// TIA Portal project "OP-TQ-01" (V13)

(* hardware
DEVICE "S7-1200 station_1"  S7-1200 Station
   slot 0: "Rack_0"  Rack  V1.0
   slot 1: "PLC_1"  CPU 1214C DC/DC/Rly  6ES7 214-1HG31-0XB0  V3.0
   slot 2: "AI 4x13BIT_1"  6ES7 231-4HD30-0XB0  V1.0
   slot 3: "AI 4x13BIT_2"  6ES7 231-4HD30-0XB0  V1.0
   slot 4: "AQ 2x14BIT_1"  6ES7 232-4HB32-0XB0  V2.0
DEVICE "HMI_1"  KP400 Comfort
   slot 0: "HMI"  HMI  6AV2 124-1DC01-0AX0  13.0.1.0
   slot 1: "HMI_RT_1"  KP400 Comfort  6AV2 124-1DC01-0AX0  13.0.1.0
   slot 5: "HMI_1.IE_CP_1"  PROFINET Interface
      slot 1: "PROFINET Interface_1"  PROFINET Interface
         slot 1: "Port_1"  Port
   slot 7: "HMI_1.MPI/DP_CP_1"  MPI/DP Interface
*)

// ===== PLC "PLC_1"  CPU 1214C DC/DC/Rly =====

VAR_GLOBAL   // PLC tag table "Default tag table"
   "System_Byte" AT %MB1 : Byte;
   "FirstScan" AT %M1.0 : Bool;
   "DiagStatusUpdate" AT %M1.1 : Bool;
   "AlwaysTRUE" AT %M1.2 : Bool;
   "AlwaysFALSE" AT %M1.3 : Bool;
   "Clock_Byte" AT %MB0 : Byte;
   "Clock_10Hz" AT %M0.0 : Bool;
   "Clock_5Hz" AT %M0.1 : Bool;
   "Clock_2.5Hz" AT %M0.2 : Bool;
   "Clock_2Hz" AT %M0.3 : Bool;
   "Clock_1.25Hz" AT %M0.4 : Bool;
   "Clock_1Hz" AT %M0.5 : Bool;
   "Clock_0.625Hz" AT %M0.6 : Bool;
   "Clock_0.5Hz" AT %M0.7 : Bool;
   "TT-006-EA" AT %IW96 : Int;
   "TT-007-EA" AT %IW98 : Int;
   "TT-008-EA" AT %IW100 : Int;
   "TT-009-EA" AT %IW102 : Int;
   "TT-010-EA" AT %IW104 : Int;
   "TT-011-EA" AT %IW106 : Int;
   "LT-009-EA" AT %IW108 : Int;
   "LT-CX-REC-EA" AT %IW110 : Int;
   "LSLL-004" AT %I0.0 : Bool;
   "TSH-004" AT %I0.1 : Bool;
   "TERMICO" AT %I0.2 : Bool;
   "RESISTENCIAS-MAN-AUTO" AT %I0.3 : Bool;
   "RESISTENCIAS-RETORNO" AT %I0.4 : Bool;
   "BOTAO-LIGA" AT %I0.5 : Bool;
   "BOTAO-DESLIGA" AT %I0.6 : Bool;
   "FALTA-DE-FASE" AT %I0.7 : Bool;
   "RESISTENCIAS-DESLIGA" AT %Q0.0 : Bool;
   "R2-DESLIGA" AT %Q0.1 : Bool;
   "CX-REC-NIVEL-H" AT %Q0.2 : Bool;
   "CX-REC-NIVEL-HH" AT %Q0.3 : Bool;
   "AlarmAnalog" AT %M13.0 : Bool;
   "REC_ALM" AT %M2.0 : Bool;
   "IW0" AT %IW0 : Word;
   "SAIDAS_DIGITAIS" AT %QW0 : Word;
   "R01A-Liga" AT %M110.0 : Bool;
   "R01B-Liga" AT %M110.1 : Bool;
   "R01C-Liga" AT %M110.2 : Bool;
   "R01D-Liga" AT %M110.3 : Bool;
   "R01E-Liga" AT %M110.4 : Bool;
   "R01F-Liga" AT %M110.5 : Bool;
   "Intlok-Resist" AT %M110.6 : Bool;
   "Tag_1" AT %MW140 : Int;
   "Tag_2" AT %MW142 : Int;
   "Tag_3" AT %MW144 : Int;
   "Tag_4" AT %M20.0 : Bool;
   "Tag_5" AT %M20.1 : Bool;
END_VAR

TYPE "Alm-Bits"
   STRUCT
      UDF : Bool;
      UDR : Bool;
      OVF : Bool;
      OVR : Bool;
      HH : Bool;
      H : Bool;
      L : Bool;
      LL : Bool;
   END_STRUCT;
END_TYPE

TYPE "SP-Temperaturas"
   STRUCT
      AuxLiga : Bool;
      ErroSP : Bool;
      "SP-MAX" : Real;
      "SP-MIN" : Real;
   END_STRUCT;
END_TYPE

// folder: 0000 - AUXILIARES

DATA_BLOCK "TIMERS"   // DB5100
{ S7_Optimized_Access := 'FALSE' }
VERSION : 0.1
   VAR
      T : Array[0..25] of IEC_TIMER;
   END_VAR
BEGIN
END_DATA_BLOCK

// folder: 0020 - ENTRADAS DIGITAIS

DATA_BLOCK "ED"   // DB20
TITLE = ESPELHO DAS ENTRADAS DIGITAIS
{ S7_Optimized_Access := 'FALSE' }
VERSION : 0.1
   VAR
      "LSLL-004" : Bool;
      "TSH-004" : Bool;
      TERMICO : Bool;
      "RESISTENCIAS-LOC-REM" : Bool;
      "RESISTENCIAS-RETORNO" : Bool;
      "BOTAO-LIGA" : Bool;
      "BOTAO-DESLIGA" : Bool;
      "FALTA-DE-FASE" : Bool;
      RESERVA_1 : Bool;
      RESERVA_2 : Bool;
      RESERVA_3 : Bool;
      RESERVA_4 : Bool;
      RESERVA_5 : Bool;
      RESERVA_6 : Bool;
      RESERVA_7 : Bool;
      RESERVA_8 : Bool;
      RESERVA : Array[2..3] of Byte;
   END_VAR
BEGIN
END_DATA_BLOCK

// folder: 0030 - SAIDAS DIGITAIS

DATA_BLOCK "SD"   // DB30
TITLE = ESPELHO DAS SAÍDAS DIGITAIS
{ S7_Optimized_Access := 'FALSE' }
VERSION : 0.1
   VAR
      "LD-RESISTENCIAS" : Bool;
      "R2-DESLIGA" : Bool;
      "CX-REC-NIVEL-H" : Bool;
      "CX-REC-NIVEL-HH" : Bool;
      RESERVA_1 : Bool;
      RESERVA_2 : Bool;
      RESERVA_3 : Bool;
      RESERVA_4 : Bool;
      RESERVA_5 : Bool;
      RESERVA_6 : Bool;
      RESERVA_7 : Bool;
      RESERVA_8 : Bool;
      RESERVA_9 : Bool;
      RESERVA_10 : Bool;
      RESERVA_11 : Bool;
      RESERVA_12 : Bool;
      RESERVA : Array[2..3] of Byte;
   END_VAR
BEGIN
END_DATA_BLOCK

// folder: 1100 - ACIONAMENTOS/RESISTENCIAS

DATA_BLOCK "R01A-R01F"   // DB1101
{ S7_Optimized_Access := 'FALSE' }
VERSION : 0.1
// stored: InstanceOfName 1110 - RESISTENCIAS
"1110 - RESISTENCIAS"
BEGIN
END_DATA_BLOCK

DATA_BLOCK "SP-TT"   // DB1110
{ S7_Optimized_Access := 'FALSE' }
VERSION : 0.1
   VAR
      "TT-006-R01A" : "SP-Temperaturas";
      "TT-007-R01B" : "SP-Temperaturas";
      "TT-008-R01C" : "SP-Temperaturas";
      "TT-009-R01D" : "SP-Temperaturas";
      "TT-010-R01E" : "SP-Temperaturas";
      "TT-011-R01F" : "SP-Temperaturas";
   END_VAR
BEGIN
END_DATA_BLOCK

// folder: 1300 - ALARMES

DATA_BLOCK "ALM"   // DB1301
{ S7_Optimized_Access := 'FALSE' }
VERSION : 0.1
   VAR
      "LSLL-004" : Bool;
      "TSH-004" : Bool;
      FaltaDeFase : Bool;
      RESERVA : Word;
   END_VAR
BEGIN
END_DATA_BLOCK

// folder: 1400 - ENTRADAS ANALOGICAS/NIVEL

DATA_BLOCK "LT-009"   // DB1417
{ S7_Optimized_Access := 'FALSE' }
VERSION : 0.1
// stored: InstanceOfName 1401 - LEITURAS ANALÓGICAS 1HAB
"1401 - LEITURAS ANALÓGICAS 1HAB"
BEGIN
END_DATA_BLOCK

DATA_BLOCK "LT-008"   // DB1418
{ S7_Optimized_Access := 'FALSE' }
VERSION : 0.1
// stored: InstanceOfName 1401 - LEITURAS ANALÓGICAS 1HAB
"1401 - LEITURAS ANALÓGICAS 1HAB"
BEGIN
END_DATA_BLOCK

// folder: 1400 - ENTRADAS ANALOGICAS/TEMPERATURA

DATA_BLOCK "TT-006-R01A"   // DB1411
{ S7_Optimized_Access := 'FALSE' }
VERSION : 0.1
// stored: InstanceOfName 1401 - LEITURAS ANALÓGICAS 1HAB
"1401 - LEITURAS ANALÓGICAS 1HAB"
BEGIN
END_DATA_BLOCK

DATA_BLOCK "TT-007-R01B"   // DB1412
{ S7_Optimized_Access := 'FALSE' }
VERSION : 0.1
// stored: InstanceOfName 1401 - LEITURAS ANALÓGICAS 1HAB
"1401 - LEITURAS ANALÓGICAS 1HAB"
BEGIN
END_DATA_BLOCK

DATA_BLOCK "TT-008-R01C"   // DB1413
{ S7_Optimized_Access := 'FALSE' }
VERSION : 0.1
// stored: InstanceOfName 1401 - LEITURAS ANALÓGICAS 1HAB
"1401 - LEITURAS ANALÓGICAS 1HAB"
BEGIN
END_DATA_BLOCK

DATA_BLOCK "TT-009-R01D"   // DB1414
{ S7_Optimized_Access := 'FALSE' }
VERSION : 0.1
// stored: InstanceOfName 1401 - LEITURAS ANALÓGICAS 1HAB
"1401 - LEITURAS ANALÓGICAS 1HAB"
BEGIN
END_DATA_BLOCK

DATA_BLOCK "TT-010-R01E"   // DB1415
{ S7_Optimized_Access := 'FALSE' }
VERSION : 0.1
// stored: InstanceOfName 1401 - LEITURAS ANALÓGICAS 1HAB
"1401 - LEITURAS ANALÓGICAS 1HAB"
BEGIN
END_DATA_BLOCK

DATA_BLOCK "TT-011-R01F"   // DB1416
{ S7_Optimized_Access := 'FALSE' }
VERSION : 0.1
// stored: InstanceOfName 1401 - LEITURAS ANALÓGICAS 1HAB
"1401 - LEITURAS ANALÓGICAS 1HAB"
BEGIN
END_DATA_BLOCK

// folder: (top level)

ORGANIZATION_BLOCK "Main"   // OB1, LAD, ProgramCycle
TITLE = "Main Program Sweep (Cycle)"
{ S7_Optimized_Access := 'FALSE' }
VERSION : 0.1
BEGIN

REGION Network 1
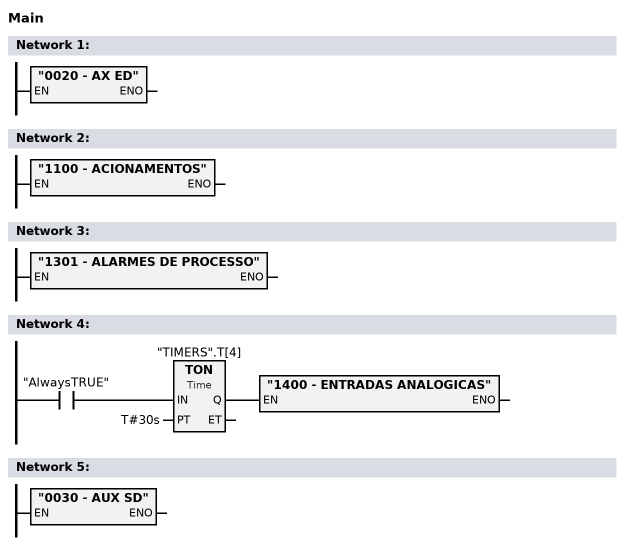
   RUNG wire#powerrail
      "0020 - AX ED"()
   END_RUNG
   // the same network as SCL:
   "0020 - AX ED"();
END_REGION

REGION Network 2
   RUNG wire#powerrail
      "1100 - ACIONAMENTOS"()
   END_RUNG
   // the same network as SCL:
   "1100 - ACIONAMENTOS"();
END_REGION

REGION Network 3
   RUNG wire#powerrail
      "1301 - ALARMES DE PROCESSO"()
   END_RUNG
   // the same network as SCL:
   "1301 - ALARMES DE PROCESSO"();
END_REGION

REGION Network 4
   "TIMERS".T[4].TON(IN := "AlwaysTRUE", PT := T#30s);
   IF "TIMERS".T[4].Q THEN "1400 - ENTRADAS ANALOGICAS"(); END_IF;
END_REGION

REGION Network 5
   RUNG wire#powerrail
      "0030 - AUX SD"()
   END_RUNG
   // the same network as SCL:
   "0030 - AUX SD"();
END_REGION
END_ORGANIZATION_BLOCK

// folder: 0020 - ENTRADAS DIGITAIS

FUNCTION "0020 - AX ED" : Void   // FC20, LAD
TITLE = ESPELHO DAS ENTRADAS DIGITAIS
{ S7_Optimized_Access := 'FALSE' }
VERSION : 0.1
BEGIN

REGION Network 1: ESPELHA AS ENTRADAS DIGITAIS DO CLP
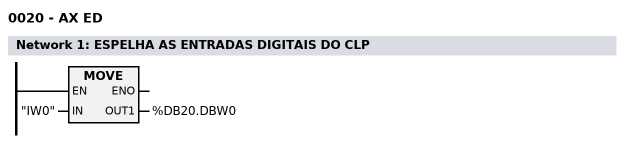
   RUNG wire#powerrail
      { S7_GenerateENO := "TRUE" } Move(in := "IW0", out1 => %DB20.DBW0)
   END_RUNG
   // the same network as SCL:
   %DB20.DBW0 := "IW0";
END_REGION
END_FUNCTION

// folder: 0030 - SAIDAS DIGITAIS

FUNCTION "0030 - AUX SD" : Void   // FC30, LAD
TITLE = ESPELHO DAS SAIDAS DIGITAIS
{ S7_Optimized_Access := 'FALSE' }
VERSION : 0.1
BEGIN

REGION Network 1: ESPELHO DAS SAIDAS DIGITAIS DAS ECP1 E ECP2
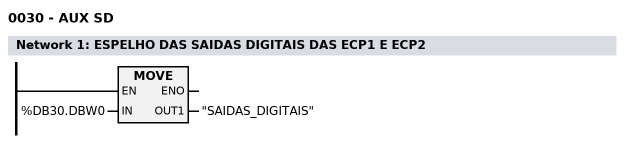
   RUNG wire#powerrail
      { S7_GenerateENO := "TRUE" } Move(in := %DB30.DBW0, out1 => "SAIDAS_DIGITAIS")
   END_RUNG
   // the same network as SCL:
   "SAIDAS_DIGITAIS" := %DB30.DBW0;
END_REGION
END_FUNCTION

// folder: 1100 - ACIONAMENTOS

FUNCTION "1100 - ACIONAMENTOS" : Void   // FC1100, LAD
TITLE = CHAMADA DOS BLOCOS DE ACIONAMENTOS DOS EQUIPAMENTOS
{ S7_Optimized_Access := 'FALSE' }
VERSION : 0.1
BEGIN

REGION Network 1: RESISTÊNCIAS R1-R6
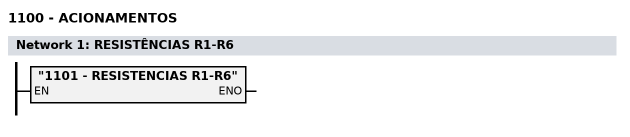
   RUNG wire#powerrail
      "1101 - RESISTENCIAS R1-R6"()
   END_RUNG
   // the same network as SCL:
   "1101 - RESISTENCIAS R1-R6"();
END_REGION
END_FUNCTION

// folder: 1100 - ACIONAMENTOS/RESISTENCIAS

FUNCTION "1101 - RESISTENCIAS R1-R6" : Void   // FC1101, LAD
TITLE = ACIONAMENTO DAS RESISTENCIAS DE AQUECIMENTO DO TQ-01
{ S7_Optimized_Access := 'FALSE' }
VERSION : 0.1
BEGIN

REGION Network 1: VERIFICA TEMPERATURA PARA LIGAR RESISTÊNCIA - R01A
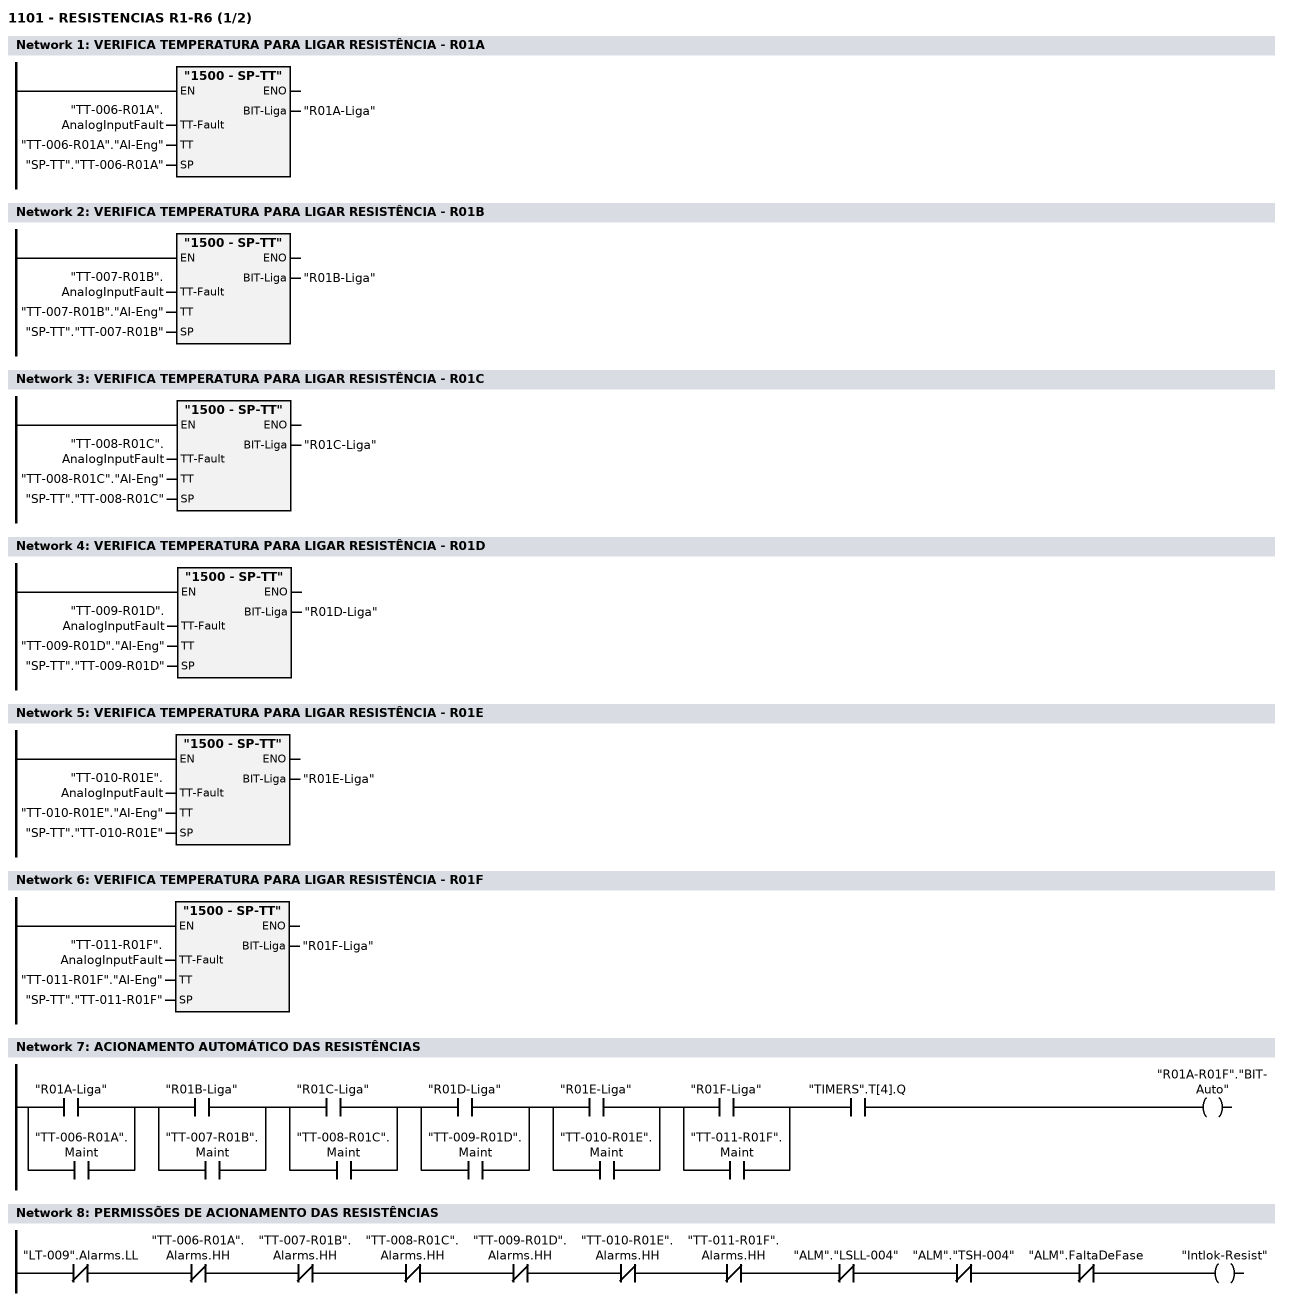
   RUNG wire#powerrail
      "1500 - SP-TT"("TT-Fault" := "TT-006-R01A".AnalogInputFault, TT := "TT-006-R01A"."AI-Eng", SP := "SP-TT"."TT-006-R01A", "BIT-Liga" => "R01A-Liga")
   END_RUNG
   // the same network as SCL:
   "1500 - SP-TT"("TT-Fault" := "TT-006-R01A".AnalogInputFault,
                  TT := "TT-006-R01A"."AI-Eng",
                  SP := "SP-TT"."TT-006-R01A",
                  "BIT-Liga" => "R01A-Liga");
END_REGION

REGION Network 2: VERIFICA TEMPERATURA PARA LIGAR RESISTÊNCIA - R01B
   RUNG wire#powerrail
      "1500 - SP-TT"("TT-Fault" := "TT-007-R01B".AnalogInputFault, TT := "TT-007-R01B"."AI-Eng", SP := "SP-TT"."TT-007-R01B", "BIT-Liga" => "R01B-Liga")
   END_RUNG
   // the same network as SCL:
   "1500 - SP-TT"("TT-Fault" := "TT-007-R01B".AnalogInputFault,
                  TT := "TT-007-R01B"."AI-Eng",
                  SP := "SP-TT"."TT-007-R01B",
                  "BIT-Liga" => "R01B-Liga");
END_REGION

REGION Network 3: VERIFICA TEMPERATURA PARA LIGAR RESISTÊNCIA - R01C
   RUNG wire#powerrail
      "1500 - SP-TT"("TT-Fault" := "TT-008-R01C".AnalogInputFault, TT := "TT-008-R01C"."AI-Eng", SP := "SP-TT"."TT-008-R01C", "BIT-Liga" => "R01C-Liga")
   END_RUNG
   // the same network as SCL:
   "1500 - SP-TT"("TT-Fault" := "TT-008-R01C".AnalogInputFault,
                  TT := "TT-008-R01C"."AI-Eng",
                  SP := "SP-TT"."TT-008-R01C",
                  "BIT-Liga" => "R01C-Liga");
END_REGION

REGION Network 4: VERIFICA TEMPERATURA PARA LIGAR RESISTÊNCIA - R01D
   RUNG wire#powerrail
      "1500 - SP-TT"("TT-Fault" := "TT-009-R01D".AnalogInputFault, TT := "TT-009-R01D"."AI-Eng", SP := "SP-TT"."TT-009-R01D", "BIT-Liga" => "R01D-Liga")
   END_RUNG
   // the same network as SCL:
   "1500 - SP-TT"("TT-Fault" := "TT-009-R01D".AnalogInputFault,
                  TT := "TT-009-R01D"."AI-Eng",
                  SP := "SP-TT"."TT-009-R01D",
                  "BIT-Liga" => "R01D-Liga");
END_REGION

REGION Network 5: VERIFICA TEMPERATURA PARA LIGAR RESISTÊNCIA - R01E
   RUNG wire#powerrail
      "1500 - SP-TT"("TT-Fault" := "TT-010-R01E".AnalogInputFault, TT := "TT-010-R01E"."AI-Eng", SP := "SP-TT"."TT-010-R01E", "BIT-Liga" => "R01E-Liga")
   END_RUNG
   // the same network as SCL:
   "1500 - SP-TT"("TT-Fault" := "TT-010-R01E".AnalogInputFault,
                  TT := "TT-010-R01E"."AI-Eng",
                  SP := "SP-TT"."TT-010-R01E",
                  "BIT-Liga" => "R01E-Liga");
END_REGION

REGION Network 6: VERIFICA TEMPERATURA PARA LIGAR RESISTÊNCIA - R01F
   RUNG wire#powerrail
      "1500 - SP-TT"("TT-Fault" := "TT-011-R01F".AnalogInputFault, TT := "TT-011-R01F"."AI-Eng", SP := "SP-TT"."TT-011-R01F", "BIT-Liga" => "R01F-Liga")
   END_RUNG
   // the same network as SCL:
   "1500 - SP-TT"("TT-Fault" := "TT-011-R01F".AnalogInputFault,
                  TT := "TT-011-R01F"."AI-Eng",
                  SP := "SP-TT"."TT-011-R01F",
                  "BIT-Liga" => "R01F-Liga");
END_REGION

REGION Network 7: ACIONAMENTO AUTOMÁTICO DAS RESISTÊNCIAS
   RUNG wire#powerrail
      Contact( "R01A-Liga" )
      wire#w1
      Contact( "R01B-Liga" )
      wire#w2
      Contact( "R01C-Liga" )
      wire#w3
      Contact( "R01D-Liga" )
      wire#w4
      Contact( "R01E-Liga" )
      wire#w5
      Contact( "R01F-Liga" )
      wire#w6
      Contact( "TIMERS".T[4].Q )
      Coil( "R01A-R01F"."BIT-Auto" )
   END_RUNG
   RUNG wire#powerrail
      Contact( "TT-006-R01A".Maint )
   END_RUNG wire#w1
   RUNG wire#w1
      Contact( "TT-007-R01B".Maint )
   END_RUNG wire#w2
   RUNG wire#w2
      Contact( "TT-008-R01C".Maint )
   END_RUNG wire#w3
   RUNG wire#w3
      Contact( "TT-009-R01D".Maint )
   END_RUNG wire#w4
   RUNG wire#w4
      Contact( "TT-010-R01E".Maint )
   END_RUNG wire#w5
   RUNG wire#w5
      Contact( "TT-011-R01F".Maint )
   END_RUNG wire#w6
   // the same network as SCL:
   "R01A-R01F"."BIT-Auto" := ("R01A-Liga" OR "TT-006-R01A".Maint) AND ("R01B-Liga" OR "TT-007-R01B".Maint) AND ("R01C-Liga" OR "TT-008-R01C".Maint) AND ("R01D-Liga" OR "TT-009-R01D".Maint) AND ("R01E-Liga" OR "TT-010-R01E".Maint) AND ("R01F-Liga" OR "TT-011-R01F".Maint) AND "TIMERS".T[4].Q;
END_REGION

REGION Network 8: PERMISSÕES DE ACIONAMENTO DAS RESISTÊNCIAS
   RUNG wire#powerrail
      I_Contact( "LT-009".Alarms.LL )
      I_Contact( "TT-006-R01A".Alarms.HH )
      I_Contact( "TT-007-R01B".Alarms.HH )
      I_Contact( "TT-008-R01C".Alarms.HH )
      I_Contact( "TT-009-R01D".Alarms.HH )
      I_Contact( "TT-010-R01E".Alarms.HH )
      I_Contact( "TT-011-R01F".Alarms.HH )
      I_Contact( "ALM"."LSLL-004" )
      I_Contact( "ALM"."TSH-004" )
      I_Contact( "ALM".FaltaDeFase )
      Coil( "Intlok-Resist" )
   END_RUNG
   // the same network as SCL:
   "Intlok-Resist" := NOT "LT-009".Alarms.LL AND NOT "TT-006-R01A".Alarms.HH AND NOT "TT-007-R01B".Alarms.HH AND NOT "TT-008-R01C".Alarms.HH AND NOT "TT-009-R01D".Alarms.HH AND NOT "TT-010-R01E".Alarms.HH AND NOT "TT-011-R01F".Alarms.HH AND NOT "ALM"."LSLL-004" AND NOT "ALM"."TSH-004" AND NOT "ALM".FaltaDeFase;
END_REGION

REGION Network 9: CHAMADA DO BLOCO PADRÃO DE ACIONAMENTO
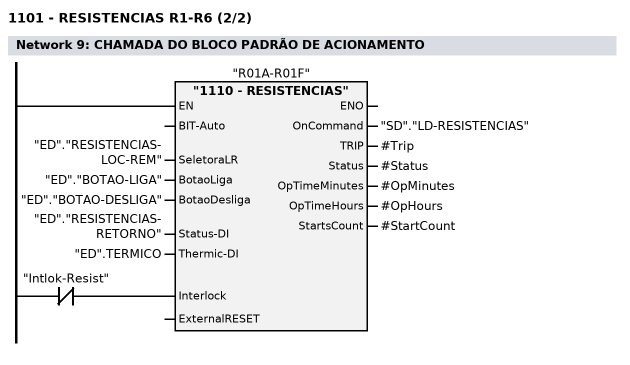
   RUNG wire#powerrail
      "R01A-R01F"(Interlock := wire#w1, "BIT-Auto" :=, SeletoraLR := "ED"."RESISTENCIAS-LOC-REM", BotaoLiga := "ED"."BOTAO-LIGA", BotaoDesliga := "ED"."BOTAO-DESLIGA", "Status-DI" := "ED"."RESISTENCIAS-RETORNO", "Thermic-DI" := "ED".TERMICO, ExternalRESET :=, OnCommand => "SD"."LD-RESISTENCIAS", TRIP => #Trip, Status => #Status, OpTimeMinutes => #OpMinutes, OpTimeHours => #OpHours, StartsCount => #StartCount)
   END_RUNG
   RUNG wire#powerrail
      I_Contact( "Intlok-Resist" )
   END_RUNG wire#w1
   // the same network as SCL:
   "R01A-R01F"(SeletoraLR := "ED"."RESISTENCIAS-LOC-REM",   // "1110 - RESISTENCIAS"
               BotaoLiga := "ED"."BOTAO-LIGA",
               BotaoDesliga := "ED"."BOTAO-DESLIGA",
               "Status-DI" := "ED"."RESISTENCIAS-RETORNO",
               "Thermic-DI" := "ED".TERMICO,
               Interlock := NOT "Intlok-Resist",
               OnCommand => "SD"."LD-RESISTENCIAS",
               TRIP => #Trip,
               Status => #Status,
               OpTimeMinutes => #OpMinutes,
               OpTimeHours => #OpHours,
               StartsCount => #StartCount);
END_REGION
END_FUNCTION

// folder: 1300 - ALARMES

FUNCTION "1301 - ALARMES DE PROCESSO" : Void   // FC1301, LAD
TITLE = ALARMES DE PROCESSO
{ S7_Optimized_Access := 'FALSE' }
VERSION : 0.1
BEGIN

REGION Network 1: CHAVE DE NÍVEL MUITO BAIXO
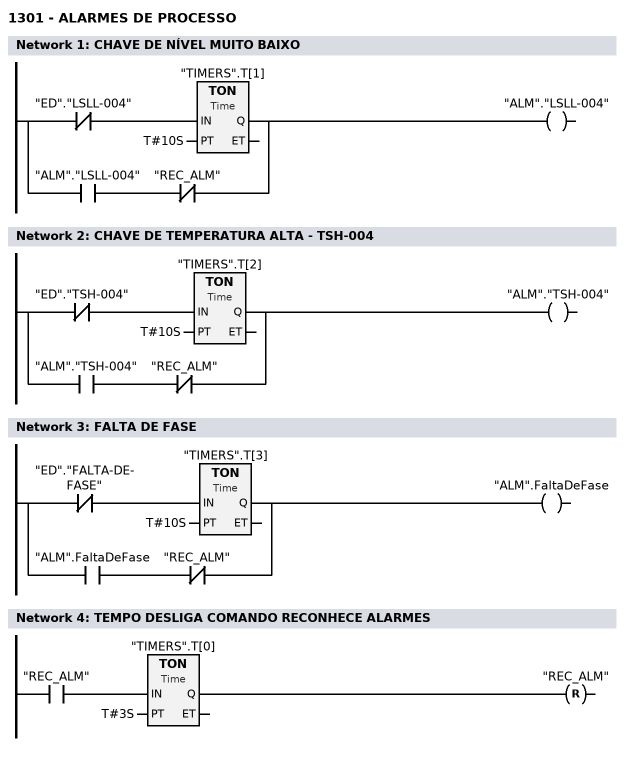
   "TIMERS".T[1].TON(IN := NOT "ED"."LSLL-004", PT := T#10S);
   "ALM"."LSLL-004" := "TIMERS".T[1].Q OR ("ALM"."LSLL-004" AND NOT "REC_ALM");
END_REGION

REGION Network 2: CHAVE DE TEMPERATURA ALTA - TSH-004
   "TIMERS".T[2].TON(IN := NOT "ED"."TSH-004", PT := T#10S);
   "ALM"."TSH-004" := "TIMERS".T[2].Q OR ("ALM"."TSH-004" AND NOT "REC_ALM");
END_REGION

REGION Network 3: FALTA DE FASE
   "TIMERS".T[3].TON(IN := NOT "ED"."FALTA-DE-FASE", PT := T#10S);
   "ALM".FaltaDeFase := "TIMERS".T[3].Q OR ("ALM".FaltaDeFase AND NOT "REC_ALM");
END_REGION

REGION Network 4: TEMPO DESLIGA COMANDO RECONHECE ALARMES
   "TIMERS".T[0].TON(IN := "REC_ALM", PT := T#3S);
   IF "TIMERS".T[0].Q THEN "REC_ALM" := FALSE; END_IF;
END_REGION
END_FUNCTION

// folder: 1400 - ENTRADAS ANALOGICAS

FUNCTION "1400 - ENTRADAS ANALOGICAS" : Void   // FC1400, LAD
{ S7_Optimized_Access := 'FALSE' }
VERSION : 0.1
BEGIN

REGION Network 1: RACK 00 - SLOT 02 EA 00 - RESISTENCIA 01A TQ-OP-01
   // ESCALONAMENTO DA ENTRADA 01 - RESISTENCIA TQ-OP-00
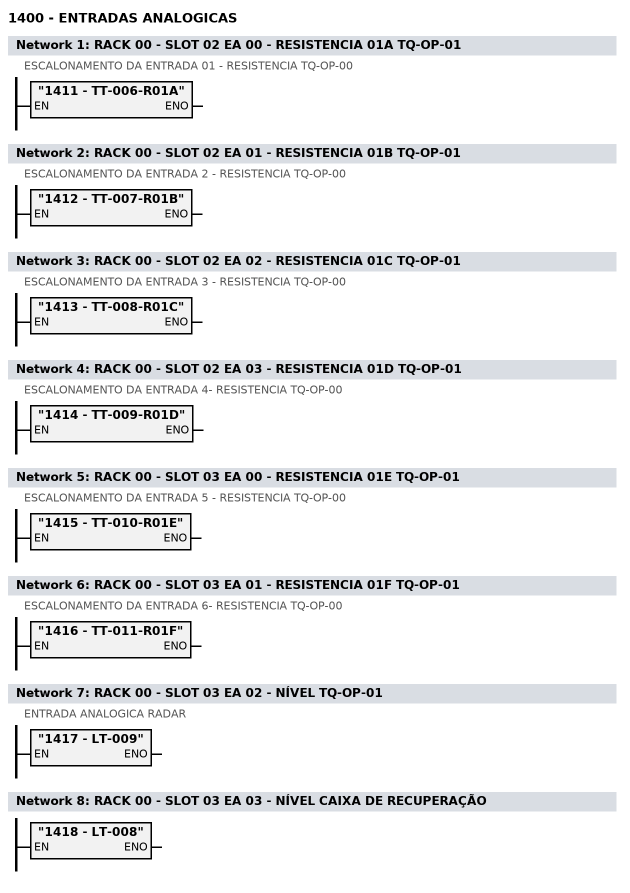
   RUNG wire#powerrail
      "1411 - TT-006-R01A"()
   END_RUNG
   // the same network as SCL:
   "1411 - TT-006-R01A"();
END_REGION

REGION Network 2: RACK 00 - SLOT 02 EA 01 - RESISTENCIA 01B TQ-OP-01
   // ESCALONAMENTO DA ENTRADA 2 - RESISTENCIA TQ-OP-00
   RUNG wire#powerrail
      "1412 - TT-007-R01B"()
   END_RUNG
   // the same network as SCL:
   "1412 - TT-007-R01B"();
END_REGION

REGION Network 3: RACK 00 - SLOT 02 EA 02 - RESISTENCIA 01C TQ-OP-01
   // ESCALONAMENTO DA ENTRADA 3 - RESISTENCIA TQ-OP-00
   RUNG wire#powerrail
      "1413 - TT-008-R01C"()
   END_RUNG
   // the same network as SCL:
   "1413 - TT-008-R01C"();
END_REGION

REGION Network 4: RACK 00 - SLOT 02 EA 03 - RESISTENCIA 01D TQ-OP-01
   // ESCALONAMENTO DA ENTRADA 4- RESISTENCIA TQ-OP-00
   RUNG wire#powerrail
      "1414 - TT-009-R01D"()
   END_RUNG
   // the same network as SCL:
   "1414 - TT-009-R01D"();
END_REGION

REGION Network 5: RACK 00 - SLOT 03 EA 00 - RESISTENCIA 01E TQ-OP-01
   // ESCALONAMENTO DA ENTRADA 5 - RESISTENCIA TQ-OP-00
   RUNG wire#powerrail
      "1415 - TT-010-R01E"()
   END_RUNG
   // the same network as SCL:
   "1415 - TT-010-R01E"();
END_REGION

REGION Network 6: RACK 00 - SLOT 03 EA 01 - RESISTENCIA 01F TQ-OP-01
   // ESCALONAMENTO DA ENTRADA 6- RESISTENCIA TQ-OP-00
   RUNG wire#powerrail
      "1416 - TT-011-R01F"()
   END_RUNG
   // the same network as SCL:
   "1416 - TT-011-R01F"();
END_REGION

REGION Network 7: RACK 00 - SLOT 03 EA 02 - NÍVEL TQ-OP-01
   // ENTRADA ANALOGICA RADAR
   RUNG wire#powerrail
      "1417 - LT-009"()
   END_RUNG
   // the same network as SCL:
   "1417 - LT-009"();
END_REGION

REGION Network 8: RACK 00 - SLOT 03 EA 03 - NÍVEL CAIXA DE RECUPERAÇÃO
   RUNG wire#powerrail
      "1418 - LT-008"()
   END_RUNG
   // the same network as SCL:
   "1418 - LT-008"();
END_REGION
END_FUNCTION

// folder: 1400 - ENTRADAS ANALOGICAS/NIVEL

FUNCTION "1417 - LT-009" : Void   // FC1417, LAD
TITLE = LT-009
{ S7_Optimized_Access := 'FALSE' }
VERSION : 0.1
BEGIN

REGION Network 1: CHAMADA DO BLOCO PADRÃO DE ENTRADAS ANALÓGICAS
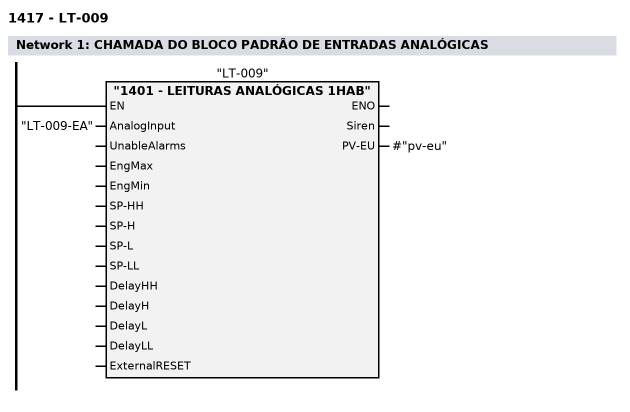
   RUNG wire#powerrail
      "LT-009"(AnalogInput := "LT-009-EA", UnableAlarms :=, EngMax :=, EngMin :=, "SP-HH" :=, "SP-H" :=, "SP-L" :=, "SP-LL" :=, DelayHH :=, DelayH :=, DelayL :=, DelayLL :=, ExternalRESET :=, Siren =>, "PV-EU" => #"pv-eu")
   END_RUNG
   // the same network as SCL:
   "LT-009"(AnalogInput := "LT-009-EA", "PV-EU" => #"pv-eu");   // "1401 - LEITURAS ANALÓGICAS 1HAB"
END_REGION
END_FUNCTION

FUNCTION "1418 - LT-008" : Void   // FC1418, LAD
TITLE = LT-CX-REC
{ S7_Optimized_Access := 'FALSE' }
VERSION : 0.1
BEGIN

REGION Network 1: CHAMADA DO BLOCO PADRÃO DE ENTRADAS ANALÓGICAS
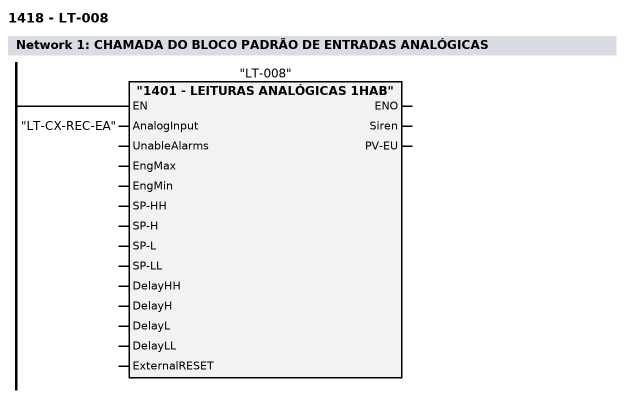
   RUNG wire#powerrail
      "LT-008"(AnalogInput := "LT-CX-REC-EA", UnableAlarms :=, EngMax :=, EngMin :=, "SP-HH" :=, "SP-H" :=, "SP-L" :=, "SP-LL" :=, DelayHH :=, DelayH :=, DelayL :=, DelayLL :=, ExternalRESET :=, Siren =>, "PV-EU" =>)
   END_RUNG
   // the same network as SCL:
   "LT-008"(AnalogInput := "LT-CX-REC-EA");   // "1401 - LEITURAS ANALÓGICAS 1HAB"
END_REGION
END_FUNCTION

// folder: 1400 - ENTRADAS ANALOGICAS/TEMPERATURA

FUNCTION "1411 - TT-006-R01A" : Void   // FC1411, LAD
TITLE = TT-006-R01A
{ S7_Optimized_Access := 'FALSE' }
VERSION : 0.1
BEGIN

REGION Network 1: CHAMADA DO BLOCO PADRÃO DE ENTRADAS ANALÓGICAS
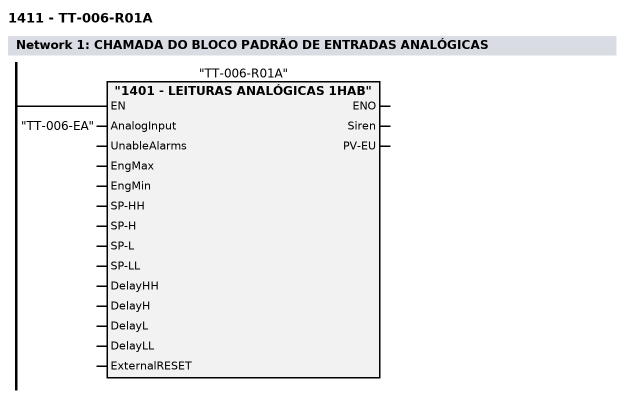
   RUNG wire#powerrail
      "TT-006-R01A"(AnalogInput := "TT-006-EA", UnableAlarms :=, EngMax :=, EngMin :=, "SP-HH" :=, "SP-H" :=, "SP-L" :=, "SP-LL" :=, DelayHH :=, DelayH :=, DelayL :=, DelayLL :=, ExternalRESET :=, Siren =>, "PV-EU" =>)
   END_RUNG
   // the same network as SCL:
   "TT-006-R01A"(AnalogInput := "TT-006-EA");   // "1401 - LEITURAS ANALÓGICAS 1HAB"
END_REGION
END_FUNCTION

FUNCTION "1412 - TT-007-R01B" : Void   // FC1412, LAD
TITLE = TT-007-R01B
{ S7_Optimized_Access := 'FALSE' }
VERSION : 0.1
BEGIN

REGION Network 1: CHAMADA DO BLOCO PADRÃO DE ENTRADAS ANALÓGICAS
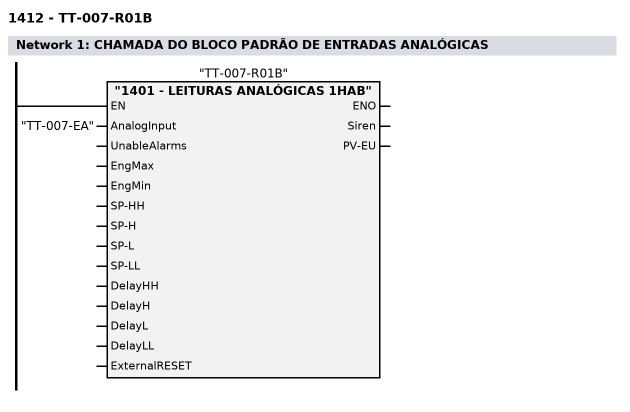
   RUNG wire#powerrail
      "TT-007-R01B"(AnalogInput := "TT-007-EA", UnableAlarms :=, EngMax :=, EngMin :=, "SP-HH" :=, "SP-H" :=, "SP-L" :=, "SP-LL" :=, DelayHH :=, DelayH :=, DelayL :=, DelayLL :=, ExternalRESET :=, Siren =>, "PV-EU" =>)
   END_RUNG
   // the same network as SCL:
   "TT-007-R01B"(AnalogInput := "TT-007-EA");   // "1401 - LEITURAS ANALÓGICAS 1HAB"
END_REGION
END_FUNCTION

FUNCTION "1413 - TT-008-R01C" : Void   // FC1413, LAD
TITLE = TT-006-R01A
{ S7_Optimized_Access := 'FALSE' }
VERSION : 0.1
BEGIN

REGION Network 1: CHAMADA DO BLOCO PADRÃO DE ENTRADAS ANALÓGICAS
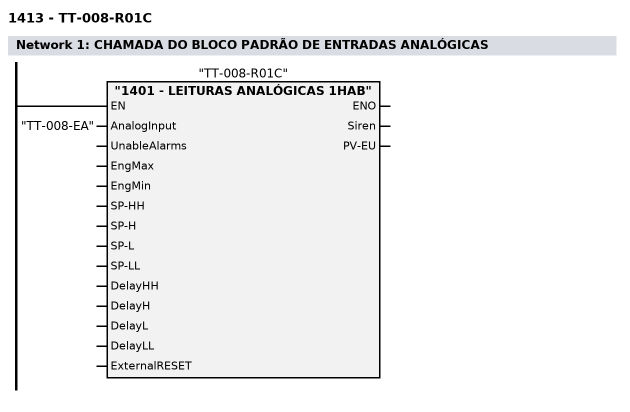
   RUNG wire#powerrail
      "TT-008-R01C"(AnalogInput := "TT-008-EA", UnableAlarms :=, EngMax :=, EngMin :=, "SP-HH" :=, "SP-H" :=, "SP-L" :=, "SP-LL" :=, DelayHH :=, DelayH :=, DelayL :=, DelayLL :=, ExternalRESET :=, Siren =>, "PV-EU" =>)
   END_RUNG
   // the same network as SCL:
   "TT-008-R01C"(AnalogInput := "TT-008-EA");   // "1401 - LEITURAS ANALÓGICAS 1HAB"
END_REGION
END_FUNCTION

FUNCTION "1414 - TT-009-R01D" : Void   // FC1414, LAD
TITLE = TT-006-R01A
{ S7_Optimized_Access := 'FALSE' }
VERSION : 0.1
BEGIN

REGION Network 1: CHAMADA DO BLOCO PADRÃO DE ENTRADAS ANALÓGICAS
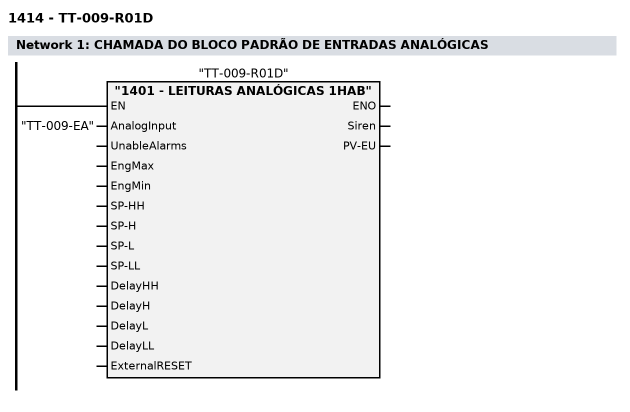
   RUNG wire#powerrail
      "TT-009-R01D"(AnalogInput := "TT-009-EA", UnableAlarms :=, EngMax :=, EngMin :=, "SP-HH" :=, "SP-H" :=, "SP-L" :=, "SP-LL" :=, DelayHH :=, DelayH :=, DelayL :=, DelayLL :=, ExternalRESET :=, Siren =>, "PV-EU" =>)
   END_RUNG
   // the same network as SCL:
   "TT-009-R01D"(AnalogInput := "TT-009-EA");   // "1401 - LEITURAS ANALÓGICAS 1HAB"
END_REGION
END_FUNCTION

FUNCTION "1415 - TT-010-R01E" : Void   // FC1415, LAD
TITLE = TT-006-R01A
{ S7_Optimized_Access := 'FALSE' }
VERSION : 0.1
BEGIN

REGION Network 1: CHAMADA DO BLOCO PADRÃO DE ENTRADAS ANALÓGICAS
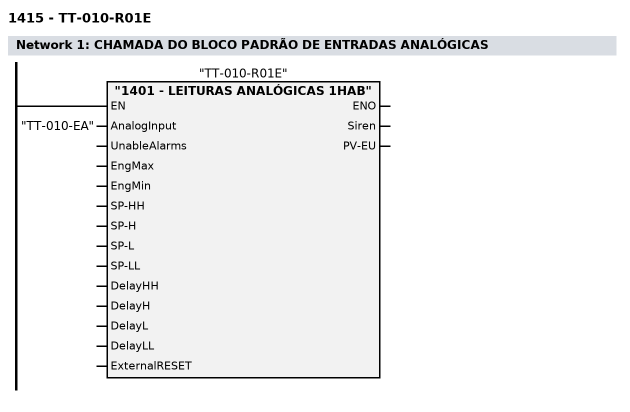
   RUNG wire#powerrail
      "TT-010-R01E"(AnalogInput := "TT-010-EA", UnableAlarms :=, EngMax :=, EngMin :=, "SP-HH" :=, "SP-H" :=, "SP-L" :=, "SP-LL" :=, DelayHH :=, DelayH :=, DelayL :=, DelayLL :=, ExternalRESET :=, Siren =>, "PV-EU" =>)
   END_RUNG
   // the same network as SCL:
   "TT-010-R01E"(AnalogInput := "TT-010-EA");   // "1401 - LEITURAS ANALÓGICAS 1HAB"
END_REGION
END_FUNCTION

FUNCTION "1416 - TT-011-R01F" : Void   // FC1416, LAD
TITLE = TT-006-R01A
{ S7_Optimized_Access := 'FALSE' }
VERSION : 0.1
BEGIN

REGION Network 1: CHAMADA DO BLOCO PADRÃO DE ENTRADAS ANALÓGICAS